// TIA Portal project "Proyecto automatizacion" (V20)

(* hardware
DEVICE "S7-1200 station_1"  S7-1200 Station
   slot 0: "Rack_0"  S7-1200 Rack  Rack  V1.0
   slot 1: "PLC_1"  CPU 1214C DC/DC/DC  6ES7 214-1AG40-0XB0  V4.7
DEVICE "HMI_1"  KTP700 Basic PN
   slot 0: "HMI_1"  KTP700 Basic PN  6AV2 123-2GB03-0AX0  17.0.0.0
   slot 1: "HMI_RT_1"  KTP700 Basic PN  6AV2 123-2GB03-0AX0  17.0.0.0
   slot 5: "HMI_1.IE_CP_1"  PROFINET Interface  17.0.0.0
      slot 1: "PROFINET Interface_1"  PROFINET Interface
         slot 1: "Port_1"  Port
*)

// ===== PLC "PLC_1"  CPU 1214C DC/DC/DC =====

VAR_GLOBAL   // PLC tag table "Default tag table"
   "1B0" AT %I0.0 : Bool;   // Sensor magnético Cilindro 1 en Home (0 mm)
   "1B1" AT %I0.1 : Bool;   // Sensor magnético Cilindro 1 en Trabajo (300 mm)
   "2B0" AT %I0.2 : Bool;   // Sensor inductivo Rotativo en Home (0°)
   "2B1" AT %I0.3 : Bool;   // Sensor inductivo Rotativo en Trabajo (90°)
   "3B0" AT %I0.4 : Bool;   // Sensor magnético Cilindro 2 en Home (0 mm)
   "3B1" AT %I0.5 : Bool;   // Sensor magnético Cilindro 2 en Trabajo (300 mm)
   "START" AT %I0.6 : Bool;   // Pulsador verde de inicio de ciclo (NA)
   "STOP" AT %I0.7 : Bool;   // Pulsador amarillo de paro a fin de ciclo (NC)
   "E_STOP" AT %I1.0 : Bool;   // Seta de Parada de Emergencia / Relé Seguridad (NC)
   "RESET" AT %I1.1 : Bool;   // Pulsador azul de rearme y homming (NA)
   "S_PESO_25KG" AT %I1.2 : Bool;   // Sensor de peso balanza en Punto A (Permiso inicio)
   "S_SACO_B" AT %I1.3 : Bool;   // Sensor presencia de saco en Punto B
   "1Y1" AT %Q0.0 : Bool;   // Solenoide Avance Cilindro 1
   "1Y0" AT %Q0.1 : Bool;   // Solenoide Retorno Cilindro 1
   "2Y1" AT %Q0.2 : Bool;   // Solenoide Giro Rotativo (Orientación 0° a 90°)
   "2Y0" AT %Q0.3 : Bool;   // Solenoide Retorno Rotativo (90° a 0°)
   "3Y1" AT %Q0.4 : Bool;   // Solenoide Avance Cilindro 2
   "3Y0" AT %Q0.5 : Bool;   // Solenoide Retorno Cilindro 2
   "H_RUN" AT %Q0.6 : Bool;   // Baliza Luz Verde (Sistema en Ciclo Automático)
   "H_ALARM" AT %Q0.7 : Bool;   // Baliza Luz Roja (Falla, Paro de Fin de Ciclo o Emergencia
   "M_RUN" AT %M0.0 : Bool;   // Relé maestro de ciclo continuo (Autorretención de START)
   "M_STOP" AT %M0.1 : Bool;   // Memoria de petición de paro ordenado a fin de ciclo
   "M_RESET" AT %M0.2 : Bool;   // Habilitación de secuencia de despeje anticolisión
   "M_ETAPA_0" AT %M1.0 : Bool;   // Estado inicial / Máquina en posición cero
   "M_ETAPA_1" AT %M1.1 : Bool;   // Avance Cilindro 1
   "M_ETAPA_2" AT %M1.2 : Bool;   // Retorno rápido Cilindro 1
   "M_ETAPA_3" AT %M1.3 : Bool;   // Giro de Actuador Rotativo a 90°
   "M_ETAPA_4" AT %M1.4 : Bool;   // Avance Cilindro 2
   "M_ETAPA_5" AT %M1.5 : Bool;   // Retorno simultáneo Rotativo y Cilindro 2
   "M_HOME_ALL" AT %M1.6 : Bool;   // Orden interna: Retraer Cilindro 1, Rotativo y CilIndro 2
   "START_HMI" AT %M0.3 : Bool;
   "STOP_HMI" AT %M0.4 : Bool;
   "RESET_HMI" AT %M0.5 : Bool;
   "Tag_1" AT %M0.6 : Bool;
END_VAR

DATA_BLOCK "DB_Alarmas"   // DB3
{ S7_Optimized_Access := 'TRUE' }
VERSION : 0.1
   VAR
      Registro_Fallos : Word;
   END_VAR
BEGIN
END_DATA_BLOCK

DATA_BLOCK "DB_Manual"   // DB4
{ S7_Optimized_Access := 'TRUE' }
VERSION : 0.1
   VAR
      Modo_Activo : Bool;
      HMI_C1_Sale : Bool;
      HMI_C1_Entra : Bool;
      HMI_C2_Sale : Bool;
      HMI_C2_Entra : Bool;
      "HMI_M_90°" : Bool;
      "HMI_M_0°" : Bool;
   END_VAR
BEGIN
END_DATA_BLOCK

// folder: System blocks/Program resources

DATA_BLOCK "IEC_Timer_0_DB"   // DB1
{ S7_Optimized_Access := 'TRUE' }
AUTHOR : Simatic
FAMILY : IEC
NAME : IEC_TMR
VERSION : 1.0
// stored: InstanceOfName IEC_TIMER
"IEC_TIMER"
BEGIN
END_DATA_BLOCK

// folder: (top level)

FUNCTION "Secuencia_Automatica" : Void   // FC1, LAD
{ S7_Optimized_Access := 'TRUE' }
VERSION : 0.1
BEGIN

REGION Network 1: Relé maestro de ciclo continuo (Autorretención de START)
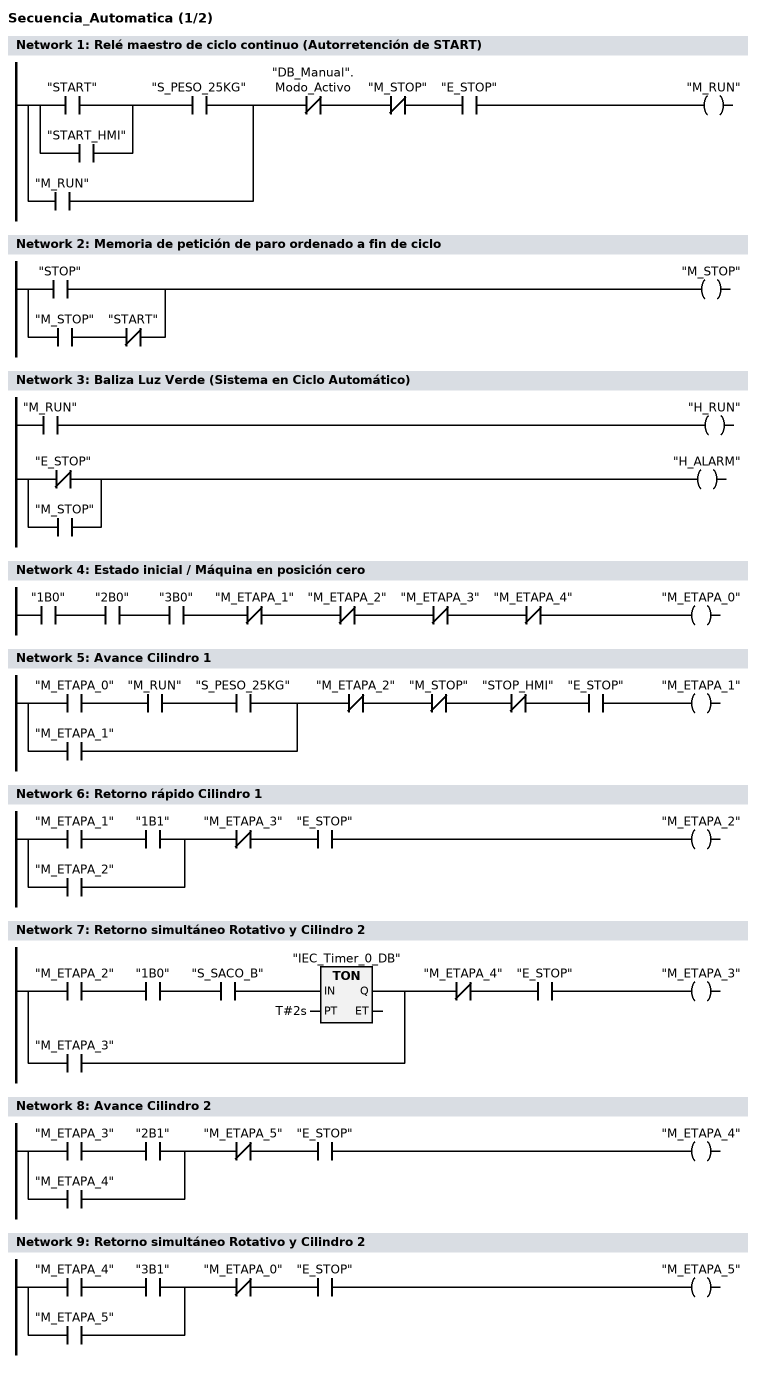
   RUNG wire#powerrail
      Contact( "START" )
      wire#w1
      Contact( "S_PESO_25KG" )
      wire#w2
      I_Contact( "DB_Manual".Modo_Activo )
      I_Contact( "M_STOP" )
      Contact( "E_STOP" )
      Coil( "M_RUN" )
   END_RUNG
   RUNG wire#powerrail
      Contact( "START_HMI" )
   END_RUNG wire#w1
   RUNG wire#powerrail
      Contact( "M_RUN" )
   END_RUNG wire#w2
   // the same network as SCL:
   "M_RUN" := ((("START" OR "START_HMI") AND "S_PESO_25KG") OR "M_RUN") AND NOT "DB_Manual".Modo_Activo AND NOT "M_STOP" AND "E_STOP";
END_REGION

REGION Network 2: Memoria de petición de paro ordenado a fin de ciclo
   RUNG wire#powerrail
      Contact( "STOP" )
      wire#w1
      Coil( "M_STOP" )
   END_RUNG
   RUNG wire#powerrail
      Contact( "M_STOP" )
      I_Contact( "START" )
   END_RUNG wire#w1
   // the same network as SCL:
   "M_STOP" := "STOP" OR ("M_STOP" AND NOT "START");
END_REGION

REGION Network 3: Baliza Luz Verde (Sistema en Ciclo Automático)
   RUNG wire#powerrail
      Contact( "M_RUN" )
      Coil( "H_RUN" )
   END_RUNG
   RUNG wire#powerrail
      I_Contact( "E_STOP" )
      wire#w1
      Coil( "H_ALARM" )
   END_RUNG
   RUNG wire#powerrail
      Contact( "M_STOP" )
   END_RUNG wire#w1
   // the same network as SCL:
   "H_RUN" := "M_RUN";
   "H_ALARM" := NOT "E_STOP" OR "M_STOP";
END_REGION

REGION Network 4: Estado inicial / Máquina en posición cero
   RUNG wire#powerrail
      Contact( "1B0" )
      Contact( "2B0" )
      Contact( "3B0" )
      I_Contact( "M_ETAPA_1" )
      I_Contact( "M_ETAPA_2" )
      I_Contact( "M_ETAPA_3" )
      I_Contact( "M_ETAPA_4" )
      Coil( "M_ETAPA_0" )
   END_RUNG
   // the same network as SCL:
   "M_ETAPA_0" := "1B0" AND "2B0" AND "3B0" AND NOT "M_ETAPA_1" AND NOT "M_ETAPA_2" AND NOT "M_ETAPA_3" AND NOT "M_ETAPA_4";
END_REGION

REGION Network 5: Avance Cilindro 1
   RUNG wire#powerrail
      Contact( "M_ETAPA_0" )
      Contact( "M_RUN" )
      Contact( "S_PESO_25KG" )
      wire#w1
      I_Contact( "M_ETAPA_2" )
      I_Contact( "M_STOP" )
      I_Contact( "STOP_HMI" )
      Contact( "E_STOP" )
      Coil( "M_ETAPA_1" )
   END_RUNG
   RUNG wire#powerrail
      Contact( "M_ETAPA_1" )
   END_RUNG wire#w1
   // the same network as SCL:
   "M_ETAPA_1" := (("M_ETAPA_0" AND "M_RUN" AND "S_PESO_25KG") OR "M_ETAPA_1") AND NOT "M_ETAPA_2" AND NOT "M_STOP" AND NOT "STOP_HMI" AND "E_STOP";
END_REGION

REGION Network 6: Retorno rápido Cilindro 1
   RUNG wire#powerrail
      Contact( "M_ETAPA_1" )
      Contact( "1B1" )
      wire#w1
      I_Contact( "M_ETAPA_3" )
      Contact( "E_STOP" )
      Coil( "M_ETAPA_2" )
   END_RUNG
   RUNG wire#powerrail
      Contact( "M_ETAPA_2" )
   END_RUNG wire#w1
   // the same network as SCL:
   "M_ETAPA_2" := (("M_ETAPA_1" AND "1B1") OR "M_ETAPA_2") AND NOT "M_ETAPA_3" AND "E_STOP";
END_REGION

REGION Network 7: Retorno simultáneo Rotativo y Cilindro 2
   "IEC_Timer_0_DB".TON(IN := "M_ETAPA_2" AND "1B0" AND "S_SACO_B", PT := T#2s);
   "M_ETAPA_3" := ("IEC_Timer_0_DB".Q OR "M_ETAPA_3") AND NOT "M_ETAPA_4" AND "E_STOP";
END_REGION

REGION Network 8: Avance Cilindro 2
   RUNG wire#powerrail
      Contact( "M_ETAPA_3" )
      Contact( "2B1" )
      wire#w1
      I_Contact( "M_ETAPA_5" )
      Contact( "E_STOP" )
      Coil( "M_ETAPA_4" )
   END_RUNG
   RUNG wire#powerrail
      Contact( "M_ETAPA_4" )
   END_RUNG wire#w1
   // the same network as SCL:
   "M_ETAPA_4" := (("M_ETAPA_3" AND "2B1") OR "M_ETAPA_4") AND NOT "M_ETAPA_5" AND "E_STOP";
END_REGION

REGION Network 9: Retorno simultáneo Rotativo y Cilindro 2
   RUNG wire#powerrail
      Contact( "M_ETAPA_4" )
      Contact( "3B1" )
      wire#w1
      I_Contact( "M_ETAPA_0" )
      Contact( "E_STOP" )
      Coil( "M_ETAPA_5" )
   END_RUNG
   RUNG wire#powerrail
      Contact( "M_ETAPA_5" )
   END_RUNG wire#w1
   // the same network as SCL:
   "M_ETAPA_5" := (("M_ETAPA_4" AND "3B1") OR "M_ETAPA_5") AND NOT "M_ETAPA_0" AND "E_STOP";
END_REGION

REGION Network 10: Orden interna: Retraer Rotativo y CilIndro 2
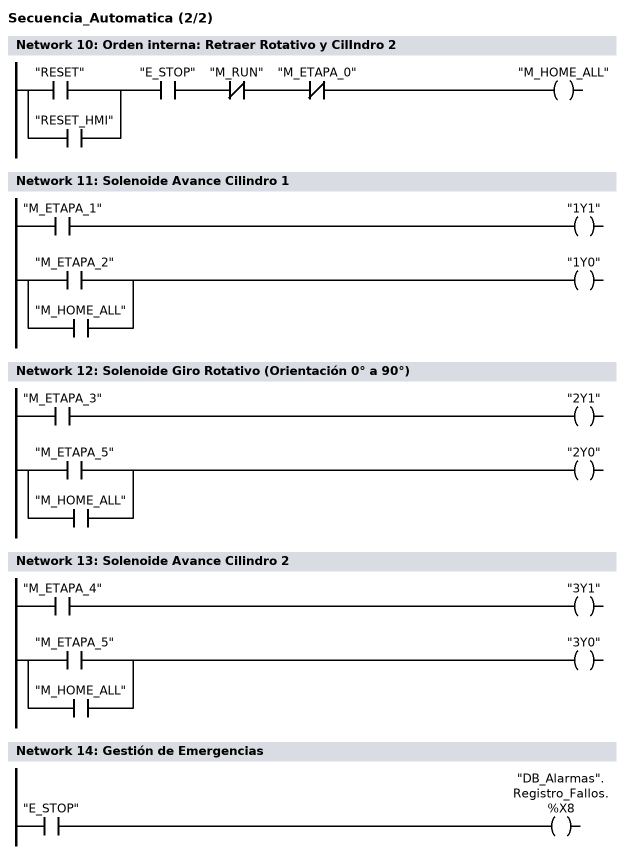
   RUNG wire#powerrail
      Contact( "RESET" )
      wire#w1
      Contact( "E_STOP" )
      I_Contact( "M_RUN" )
      I_Contact( "M_ETAPA_0" )
      Coil( "M_HOME_ALL" )
   END_RUNG
   RUNG wire#powerrail
      Contact( "RESET_HMI" )
   END_RUNG wire#w1
   // the same network as SCL:
   "M_HOME_ALL" := ("RESET" OR "RESET_HMI") AND "E_STOP" AND NOT "M_RUN" AND NOT "M_ETAPA_0";
END_REGION

REGION Network 11: Solenoide Avance Cilindro 1
   RUNG wire#powerrail
      Contact( "M_ETAPA_1" )
      Coil( "1Y1" )
   END_RUNG
   RUNG wire#powerrail
      Contact( "M_ETAPA_2" )
      wire#w1
      Coil( "1Y0" )
   END_RUNG
   RUNG wire#powerrail
      Contact( "M_HOME_ALL" )
   END_RUNG wire#w1
   // the same network as SCL:
   "1Y1" := "M_ETAPA_1";
   "1Y0" := "M_ETAPA_2" OR "M_HOME_ALL";
END_REGION

REGION Network 12: Solenoide Giro Rotativo (Orientación 0° a 90°)
   RUNG wire#powerrail
      Contact( "M_ETAPA_3" )
      Coil( "2Y1" )
   END_RUNG
   RUNG wire#powerrail
      Contact( "M_ETAPA_5" )
      wire#w1
      Coil( "2Y0" )
   END_RUNG
   RUNG wire#powerrail
      Contact( "M_HOME_ALL" )
   END_RUNG wire#w1
   // the same network as SCL:
   "2Y1" := "M_ETAPA_3";
   "2Y0" := "M_ETAPA_5" OR "M_HOME_ALL";
END_REGION

REGION Network 13: Solenoide Avance Cilindro 2
   RUNG wire#powerrail
      Contact( "M_ETAPA_4" )
      Coil( "3Y1" )
   END_RUNG
   RUNG wire#powerrail
      Contact( "M_ETAPA_5" )
      wire#w1
      Coil( "3Y0" )
   END_RUNG
   RUNG wire#powerrail
      Contact( "M_HOME_ALL" )
   END_RUNG wire#w1
   // the same network as SCL:
   "3Y1" := "M_ETAPA_4";
   "3Y0" := "M_ETAPA_5" OR "M_HOME_ALL";
END_REGION

REGION Network 14: Gestión de Emergencias
   RUNG wire#powerrail
      Contact( "E_STOP" )
      Coil( "DB_Alarmas".Registro_Fallos.%X8 )
   END_RUNG
   // the same network as SCL:
   "DB_Alarmas".Registro_Fallos.%X8 := "E_STOP";
END_REGION
END_FUNCTION

FUNCTION "FC_Control_Manual" : Void   // FC2, LAD
{ S7_Optimized_Access := 'TRUE' }
VERSION : 0.1
BEGIN

REGION Network 1: Solenoide Salida Cilindro 1
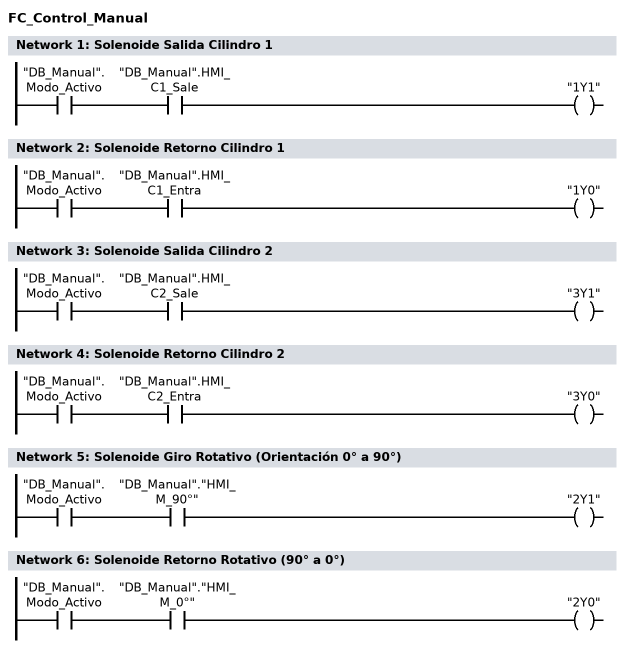
   RUNG wire#powerrail
      Contact( "DB_Manual".Modo_Activo )
      Contact( "DB_Manual".HMI_C1_Sale )
      Coil( "1Y1" )
   END_RUNG
   // the same network as SCL:
   "1Y1" := "DB_Manual".Modo_Activo AND "DB_Manual".HMI_C1_Sale;
END_REGION

REGION Network 2: Solenoide Retorno Cilindro 1
   RUNG wire#powerrail
      Contact( "DB_Manual".Modo_Activo )
      Contact( "DB_Manual".HMI_C1_Entra )
      Coil( "1Y0" )
   END_RUNG
   // the same network as SCL:
   "1Y0" := "DB_Manual".Modo_Activo AND "DB_Manual".HMI_C1_Entra;
END_REGION

REGION Network 3: Solenoide Salida Cilindro 2
   RUNG wire#powerrail
      Contact( "DB_Manual".Modo_Activo )
      Contact( "DB_Manual".HMI_C2_Sale )
      Coil( "3Y1" )
   END_RUNG
   // the same network as SCL:
   "3Y1" := "DB_Manual".Modo_Activo AND "DB_Manual".HMI_C2_Sale;
END_REGION

REGION Network 4: Solenoide Retorno Cilindro 2
   RUNG wire#powerrail
      Contact( "DB_Manual".Modo_Activo )
      Contact( "DB_Manual".HMI_C2_Entra )
      Coil( "3Y0" )
   END_RUNG
   // the same network as SCL:
   "3Y0" := "DB_Manual".Modo_Activo AND "DB_Manual".HMI_C2_Entra;
END_REGION

REGION Network 5: Solenoide Giro Rotativo (Orientación 0° a 90°)
   RUNG wire#powerrail
      Contact( "DB_Manual".Modo_Activo )
      Contact( "DB_Manual"."HMI_M_90°" )
      Coil( "2Y1" )
   END_RUNG
   // the same network as SCL:
   "2Y1" := "DB_Manual".Modo_Activo AND "DB_Manual"."HMI_M_90°";
END_REGION

REGION Network 6: Solenoide Retorno Rotativo (90° a 0°)
   RUNG wire#powerrail
      Contact( "DB_Manual".Modo_Activo )
      Contact( "DB_Manual"."HMI_M_0°" )
      Coil( "2Y0" )
   END_RUNG
   // the same network as SCL:
   "2Y0" := "DB_Manual".Modo_Activo AND "DB_Manual"."HMI_M_0°";
END_REGION
END_FUNCTION

ORGANIZATION_BLOCK "Main"   // OB1, LAD, ProgramCycle
TITLE = "Main Program Sweep (Cycle)"
{ S7_Optimized_Access := 'TRUE' }
VERSION : 0.1
   VAR_INPUT
      Initial_Call : Bool;   // Initial call of this OB
      Remanence : Bool;   // =True, if remanent data are available
   END_VAR
BEGIN

REGION Network 1
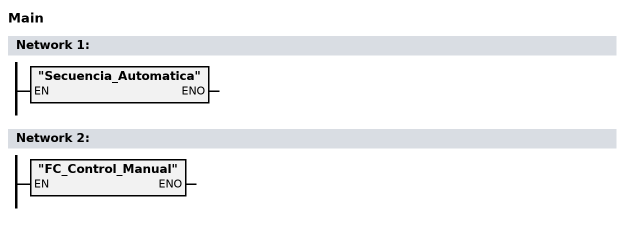
   RUNG wire#powerrail
      "Secuencia_Automatica"()
   END_RUNG
   // the same network as SCL:
   "Secuencia_Automatica"();
END_REGION

REGION Network 2
   RUNG wire#powerrail
      "FC_Control_Manual"()
   END_RUNG
   // the same network as SCL:
   "FC_Control_Manual"();
END_REGION
END_ORGANIZATION_BLOCK

(* ===== HMI "HMI_RT_1" =====
system functions are stored by id; their names below are inferred from use
connection "HMI_Connection_1": ETHERNET, SMART_S7_1200_OMS

HMI tags "Default tag table"
   "Tag_ScreenNumber" : UInt, internal
   "START_HMI" : Bool = PLC START_HMI AT %M0.3, 1 s
   "STOP_HMI" : Bool = PLC STOP_HMI AT %M0.4, 1 s
   "RESET_HMI" : Bool = PLC RESET_HMI AT %M0.5, 1 s
   "H_RUN" : Bool = PLC H_RUN AT %Q0.6, 1 s
   "H_ALARM" : Bool = PLC H_ALARM AT %Q0.7, 1 s
   "S_PESO_25KG" : Bool = PLC S_PESO_25KG AT %I1.2, 1 s
   "1B1" : Bool = PLC 1B1 AT %I0.1, 1 s
   "3B1" : Bool = PLC 3B1 AT %I0.5, 1 s
   "2B1" : Bool = PLC 2B1 AT %I0.3, 1 s
   "S_SACO_B" : Bool = PLC S_SACO_B AT %I1.3, 1 s
   "DB_Alarmas_Registro_Fallos" : Word = PLC DB_Alarmas.Registro_Fallos, 1 s
   "DB_Manual_Modo_Activo" : Bool = PLC DB_Manual.Modo_Activo, 1 s
   "DB_Manual_HMI_C1_Sale" : Bool = PLC DB_Manual.HMI_C1_Sale, 1 s
   "DB_Manual_HMI_C1_Entra" : Bool = PLC DB_Manual.HMI_C1_Entra, 1 s
   "DB_Manual_HMI_C2_Sale" : Bool = PLC DB_Manual.HMI_C2_Sale, 1 s
   "DB_Manual_HMI_C2_Entra" : Bool = PLC DB_Manual.HMI_C2_Entra, 1 s
   "DB_Manual_HMI_M_0°" : Bool = PLC DB_Manual.HMI_M_0°, 1 s
   "DB_Manual_HMI_M_90°" : Bool = PLC DB_Manual.HMI_M_90°, 1 s

discrete alarms
   1: '¡PARADA DE EMERGENCIA ACCIONADA!', class Errors, trigger "DB_Alarmas_Registro_Fallos" bit 0

Template "Template_1" 800x480
   Button "Exit" at 714,429 size 71x50; TextOff 'Exit'; PictureOff "ExitRuntime_KTP700_Basic_PN_TR"; PictureOn "ExitRuntime_KTP700_Basic_PN_TR"
      on Release: StopRuntime(0)
   Button "Start screen" at 14,429 size 71x50; TextOff 'Start screen'; PictureOff "NavigateHome_KTP700_Basic_PN_TR"; PictureOn "NavigateHome_KTP700_Basic_PN_TR"
      on Release: ActivateScreen("Principal", 0)
   SymbolicIOField "Symbolic_IO_Field_Screen" at 93,9 size 600x33; TextOff '0'; TextOn '1'; TextList "TextList_ScreenNames"
      ProcessValue <- "Tag_ScreenNumber"
      on Change: ActivateScreenByNumber("Tag_ScreenNumber", 0)
   DateTimeField "HmiScreenItemData" at 695,25 size 105x25
   DateTimeField "HmiScreenItemData_1" at 695,0 size 105x25
   GraphicView "Logo" at 0,0 size 91x51; Picture "Logo of HMI_1"
   TextField "Template_Text field_1" at 8,8 size 43x23; Text 'Text'
   Group "Group" at 114,429 size 71x50
   Button "Template_Button_5" at 114,429 size 71x50; TextOff 'Text'
      on Click: ActivateScreen("Modo_Manual", 0)
   TextField "Template_Text field_2" at 133,439 size 29x37; Text 'M'

screen "Principal" 800x480, template "Template_1"
   on GenerateScreen: SetTag("Tag_ScreenNumber", 1)
   Button "Button_1" at 12,381 size 96x32; TextOff 'START'
      on Press: SetBit("START_HMI")
      on Release: ResetBit("START_HMI")
      Appearance <- "START_HMI"
   Button "Button_2" at 124,381 size 96x32; TextOff 'STOP'
      Appearance <- "STOP_HMI"
      on Click: InvertBit("STOP_HMI")
   Button "Button_3" at 235,381 size 96x32; TextOff 'RESET'
      Appearance <- "RESET_HMI"
      on Press: SetBit("RESET_HMI")
      on Release: ResetBit("RESET_HMI")
   Circle "Circle_1" at 483,346 size 48x48
      Appearance <- "H_RUN"
   Circle "Circle_2" at 688,346 size 48x48
      Appearance <- "H_ALARM"
   TextField "Text field_1" at 458,396 size 105x23; Text 'EN MARCHA'
   TextField "Text field_2" at 646,396 size 142x23; Text 'ALARMA E-STOP'
   Rectangle "Bolsa gelatina 25 KG" at 494,177 size 91x154
      Visibility <- "S_PESO_25KG"
   Circle "Circle_3" at 319,183 size 98x98
      Visibility <- "2B1"
   Group "Group_1" at 129,129 size 135x85
   Group "Group_2" at 130,265 size 135x85
   Group "Group_3" at 108,265 size 69x85
   Group "Group" at 108,129 size 69x85
   Group "Group_4" at 319,183 size 98x98; Picture "Graphic_2"
   TextField "Text field_4" at 27,115 size 102x23; Text 'CILINDRO 1'
   TextField "Text field_5" at 28,258 size 102x23; Text 'CILINDRO 2'
   TextField "Text field_6" at 274,288 size 192x23; Text 'ACTUADOR ROTATIVO'
   TextField "Text field_7" at 464,148 size 163x23; Text 'BOLSA POSICION A'
      Visibility <- "S_PESO_25KG"
   TextField "Text field_8" at 465,148 size 162x23; Text 'BOLSA POSICION B'
      Visibility <- "S_SACO_B"
   Rectangle "Bolsa gelatina 25 KG_1" at 494,177 size 91x154
      Visibility <- "S_SACO_B"
   TextField "Text field_9" at 176,73 size 485x23; Text 'SISTEMA AUTOMÁTICO - TRANSFERENCIA POST LLENADO'
   AlarmView "Alarm view_1" at 595,183 size 197x149
      Visibility <- "DB_Alarmas_Registro_Fallos"
   Switch "Switch_1" at 361,381 size 64x32; CaptionText 'Switch'; TextOff 'OFF'; TextOn 'ON'
      ProcessValue <- "DB_Manual_Modo_Activo"
   TextField "Text field_10" at 335,358 size 131x23; Text 'MODO MANUAL'
   Circle "Circle_5" at 579,346 size 48x48
      Appearance <- "DB_Manual_Modo_Activo"
   TextField "Text field_3" at 566,395 size 76x23; Text 'MANUAL'
   Rectangle "Rectangle_2" at 108,164 size 54x19
      Visibility <- "1B1"
   Rectangle "Rectangle_3" at 153,129 size 24x85
      Visibility <- "1B1"
   Rectangle "Rectangle_5" at 129,164 size 119x19
      Visibility <- "1B1"
      Appearance <- "1B1"
   Rectangle "Rectangle_6" at 240,129 size 24x85
      Visibility <- "1B1"
      Appearance <- "1B1"
   Rectangle "Rectangle_7" at 130,300 size 119x19
      Visibility <- "3B1"
      Appearance <- "3B1"
   Rectangle "Rectangle_8" at 241,265 size 24x85
      Appearance <- "3B1"
      Visibility <- "3B1"
   Rectangle "Rectangle_9" at 108,300 size 54x19
      Visibility <- "3B1"
   Rectangle "Rectangle_10" at 153,265 size 24x85
      Visibility <- "3B1"
   GraphicView "Graphic view_2" at 342,208 size 52x52; Picture "Graphic_2"
      Visibility <- "2B1"
      Appearance <- "2B1"

screen "Root screen_1" 800x480, template "Template_1"
   on GenerateScreen: SetTag("Tag_ScreenNumber", 1)
   Button "Button_1" at 12,381 size 96x32; TextOff 'START'
      on Click: SetBit("START_HMI")
   Button "Button_2" at 119,381 size 96x32; TextOff 'STOP'
      on Click: SetBit("STOP_HMI")
   Button "Button_3" at 235,381 size 96x32; TextOff 'RESET'
      on Click: SetBit("RESET_HMI")
   Circle "Circle_1" at 548,346 size 48x48
      Appearance <- "H_RUN"
   Circle "Circle_2" at 681,346 size 48x48
      Appearance <- "H_ALARM"
   TextField "Text field_1" at 519,396 size 105x23; Text 'EN MARCHA'
   TextField "Text field_2" at 639,396 size 142x23; Text 'ALARMA E-STOP'
   Rectangle "Bolsa gelatina 25 KG" at 580,145 size 91x154
      Visibility <- "S_PESO_25KG"
   Circle "Circle_3" at 270,211 size 70x70
      Visibility <- "2B1"
   Group "Group_1" at 133,102 size 61x93
   Group "Group_2" at 70,216 size 99x62
   Group "Group_3" at 54,216 size 57x68
   Group "Group" at 134,92 size 60x48
   TextField "Text field_3" at 8,8 size 43x23; Text 'Text'
   TextField "Text field_4" at 184,53 size 102x23; Text 'CILINDRO 1'
   TextField "Text field_5" at 17,290 size 102x23; Text 'CILINDRO 2'
   TextField "Text field_6" at 225,290 size 162x23; Text 'PLATO GIRATORIO'
   TextField "Text field_7" at 552,111 size 163x23; Text 'BOLSA POSICION A'
      Visibility <- "S_PESO_25KG"
   TextField "Text field_8" at 541,92 size 162x23; Text 'BOLSA POSICION B'
      Visibility <- "S_SACO_B"
   Rectangle "Bolsa gelatina 25 KG_1" at 580,145 size 91x154
      Visibility <- "S_SACO_B"
   Group "Group_4" at 270,211 size 73x73; Picture "Graphic_2"
   Rectangle "Rectangle_2" at 156,92 size 13x38
      Visibility <- "1B1"
   Rectangle "Rectangle_3" at 134,123 size 60x17
      Visibility <- "1B1"
   Rectangle "Rectangle_5" at 155,102 size 14x82
      Visibility <- "1B1"
      Appearance <- "1B1"
   Rectangle "Rectangle_6" at 133,178 size 61x17
      Visibility <- "1B1"
      Appearance <- "1B1"
   Rectangle "Rectangle_7" at 70,242 size 87x14
      Visibility <- "3B1"
      Appearance <- "3B1"
   Rectangle "Rectangle_8" at 151,216 size 18x62
      Appearance <- "3B1"
      Visibility <- "3B1"
   Rectangle "Rectangle_9" at 54,244 size 45x15
      Visibility <- "3B1"
   Rectangle "Rectangle_10" at 91,216 size 20x68
      Visibility <- "3B1"
   GraphicView "Graphic view_2" at 283,224 size 49x51; Picture "Graphic_2"
      Visibility <- "2B1"
      Appearance <- "2B1"

screen "Modo_Manual" 800x480, template "Template_1"
   Rectangle "Rectangle_5" at 129,164 size 119x19
      Visibility <- "DB_Manual_HMI_C1_Sale"
      Appearance <- "DB_Manual_HMI_C1_Sale"
   Rectangle "Rectangle_6" at 240,129 size 24x85
      Visibility <- "DB_Manual_HMI_C1_Sale"
      Appearance <- "DB_Manual_HMI_C1_Sale"
   Rectangle "Rectangle_7" at 130,300 size 119x19
      Appearance <- "DB_Manual_HMI_C2_Sale"
      Visibility <- "DB_Manual_HMI_C2_Sale"
   Rectangle "Rectangle_8" at 241,265 size 24x85
      Appearance <- "DB_Manual_HMI_C2_Sale"
      Visibility <- "DB_Manual_HMI_C2_Sale"
   Rectangle "Rectangle_9" at 108,300 size 54x19
      Visibility <- "DB_Manual_HMI_C2_Sale"
   Rectangle "Rectangle_10" at 153,265 size 24x85
      Visibility <- "DB_Manual_HMI_C2_Sale"
   Rectangle "Rectangle_2" at 108,164 size 54x19
      Visibility <- "DB_Manual_HMI_C1_Sale"
   Rectangle "Rectangle_3" at 153,129 size 24x85
      Visibility <- "DB_Manual_HMI_C1_Sale"
   GraphicView "Graphic view_2" at 633,196 size 52x52; Picture "Graphic_2"
      Appearance <- "DB_Manual_HMI_M_90°"
      Visibility <- "DB_Manual_HMI_M_90°"
   Button "Button_1" at 12,381 size 96x32; TextOff 'START'
      on Press: SetBit("START_HMI")
      on Release: ResetBit("START_HMI")
      Appearance <- "START_HMI"
   Button "Button_2" at 124,381 size 96x32; TextOff 'STOP'
      on Click: InvertBit("STOP_HMI")
      Appearance <- "STOP_HMI"
   Button "Button_3" at 235,381 size 96x32; TextOff 'RESET'
      on Press: SetBit("RESET_HMI")
      on Release: ResetBit("RESET_HMI")
      Appearance <- "RESET_HMI"
   Circle "Circle_1" at 490,346 size 48x48
      Appearance <- "H_RUN"
   Circle "Circle_2" at 689,346 size 48x48
      Appearance <- "H_ALARM"
   TextField "Text field_1" at 454,394 size 105x23; Text 'EN MARCHA'
   TextField "Text field_2" at 647,396 size 142x23; Text 'ALARMA E-STOP'
   Circle "Circle_3" at 610,171 size 98x98
      Visibility <- "2B1"
   Group "Group_1" at 129,129 size 135x85
   Group "Group_2" at 130,265 size 135x85
   Group "Group_3" at 108,265 size 69x85
   Group "Group" at 108,129 size 69x85
   Group "Group_4" at 610,171 size 98x98; Picture "Graphic_2"
   TextField "Text field_4" at 27,115 size 102x23; Text 'CILINDRO 1'
   TextField "Text field_5" at 28,258 size 102x23; Text 'CILINDRO 2'
   TextField "Text field_6" at 565,276 size 192x23; Text 'ACTUADOR ROTATIVO'
   TextField "Text field_9" at 168,62 size 430x23; Text 'SISTEMA Manual - TRANSFERENCIA POST LLENADO'
   Switch "Switch_1" at 361,381 size 64x32; CaptionText 'Switch'; TextOff 'OFF'; TextOn 'ON'
      ProcessValue <- "DB_Manual_Modo_Activo"
   TextField "Text field_10" at 335,358 size 131x23; Text 'MODO MANUAL'
   Button "Button_4" at 555,131 size 96x32; TextOff '0°'
      on Press: SetBit("DB_Manual_HMI_M_0°")
      on Release: ResetBit("DB_Manual_HMI_M_0°")
   Button "Button_5" at 684,131 size 96x32; TextOff '90°'
      on Press: SetBit("DB_Manual_HMI_M_90°")
      on Release: ResetBit("DB_Manual_HMI_M_90°")
   Button "Button_6" at 291,119 size 96x32; TextOff 'C1 +'
      on Press: SetBit("DB_Manual_HMI_C1_Sale")
      on Release: ResetBit("DB_Manual_HMI_C1_Sale")
   Button "Button_7" at 411,119 size 96x32; TextOff 'C1 -'
      on Press: SetBit("DB_Manual_HMI_C1_Entra")
      on Release: ResetBit("DB_Manual_HMI_C1_Entra")
   Button "Button_8" at 291,244 size 96x32; TextOff 'C2 +'
      on Press: SetBit("DB_Manual_HMI_C2_Sale")
      on Release: ResetBit("DB_Manual_HMI_C2_Sale")
   Button "Button_9" at 411,244 size 96x32; TextOff 'C2 -'
      on Press: SetBit("DB_Manual_HMI_C2_Entra")
      on Release: ResetBit("DB_Manual_HMI_C2_Entra")
   TextField "Text field_3" at 567,396 size 76x23; Text 'MANUAL'
   Circle "Circle_5" at 579,346 size 48x48
      Appearance <- "DB_Manual_Modo_Activo"
*)